
screen "EPROC-ALTAMS050" 1280x800, template "Plantilla-Alta-Sec"
   Button "Botón_3" at 467,294 size 40x38; TextOff 'Text'; PictureOff "x"
      on Click: function_efd93a16()
   Button "Botón_4" at 411,540 size 96x35; TextOff 'Hecho'; Authorization "Administración de usuarios"
      on Press: SetTag("Varios_UltimoMantMS050", "HorasSecAlta_HMMS050")
   TextField "Campo de texto_6" at 37,450 size 326x27; Text 'Tiempo de funcionamiento acumulado'
   TextField "Campo de texto_4" at 37,510 size 201x27; Text 'Próximo mantenimiento'
   IOField "Campo ES_7" at 25,475 size 173x35; Authorization "Administración de usuarios"; FormatPattern 999999999; Unit  hs
      ProcessValue <- "HorasSecAlta_HMMS050"
      Appearance <- "LimiteMantMS050"
   IOField "Campo ES_1" at 205,475 size 80x35; Authorization "Administración de usuarios"; FormatPattern 99; Unit  min
      ProcessValue <- "HorasSecAlta_MMMS050"
   IOField "Campo ES_2" at 25,535 size 173x35; FormatPattern 999999999; Unit  hs
      ProcessValue <- "ProxMantMS050"
      Appearance <- "LimiteMantMS050"
   GraphicIOField "Campo ES gráfico_3" at 21,434 size 511x6; PictureList "Indicador"
      ProcessValue <- "AnimaMS050"
   TextField "Campo de texto_3" at 46,356 size 89x39; Text 'ABC 1'
   SymbolicIOField "Campo ES simbólico_3" at 48,392 size 242x21; TextOff '0'; TextOn '1'; TextList "EstadoMotor"
      ProcessValue <- "AnimaMS050"
   Switch "Interruptor_8" at 205,359 size 29x29; TextOn '1'; TextOff '0'; CaptionText 'Switch'; PictureOff "A2"; Authorization "Operación"; PictureOn "A"
      ProcessValue <- "AutoMS050"
      Visibility <- "MantMS050"
   ScreenModuleView "Faceplate_2_4" at 274,346 size 244x69
      Guid_{11997190-23979} <- "HabilitaciónMS050"
      Guid_{11997190-37146} <- "Enc1MS050"
      Guid_{11997190-23983} <- "ParadaMS050"
      Guid_{11997190-23981} <- "MarchaMS050"
      Guid_{11997190-37150} <- "Enc2MS050"
      Guid_{11997190-23976} <- "DeshabilitaciónMS050"
      Guid_{11997190-23985} <- "AnimaMenuMS050"

screen "EPROC-ALTAMS051" 1280x800, template "Plantilla-Alta-Sec"
   Button "Botón_3" at 467,294 size 40x38; TextOff 'Text'; PictureOff "x"
      on Click: function_efd93a16()
   Button "Botón_4" at 411,540 size 96x35; TextOff 'Hecho'; Authorization "Administración de usuarios"
      on Press: SetTag("Varios_UltimoMantMS051", "HorasSecAlta_HMMS051")
   TextField "Campo de texto_6" at 37,450 size 326x27; Text 'Tiempo de funcionamiento acumulado'
   TextField "Campo de texto_4" at 37,510 size 201x27; Text 'Próximo mantenimiento'
   IOField "Campo ES_7" at 25,475 size 173x35; Authorization "Administración de usuarios"; FormatPattern 999999999; Unit  hs
      ProcessValue <- "HorasSecAlta_HMMS051"
      Appearance <- "LimiteMantMS051"
   IOField "Campo ES_1" at 205,475 size 80x35; Authorization "Administración de usuarios"; FormatPattern 99; Unit  min
      ProcessValue <- "HorasSecAlta_MMMS051"
   IOField "Campo ES_2" at 25,535 size 173x35; FormatPattern 999999999; Unit  hs
      ProcessValue <- "ProxMantMS051"
      Appearance <- "LimiteMantMS051"
   GraphicIOField "Campo ES gráfico_9" at 21,434 size 511x6; PictureList "Indicador"
      ProcessValue <- "AnimaMS051"
   TextField "Campo de texto_1" at 46,356 size 89x39; Text 'ABC 3'
   SymbolicIOField "Campo ES simbólico_9" at 48,392 size 242x21; TextOff '0'; TextOn '1'; TextList "EstadoMotor"
      ProcessValue <- "AnimaMS051"
   Switch "Interruptor_5" at 211,363 size 29x29; TextOn '1'; TextOff '0'; CaptionText 'Switch'; PictureOff "A2"; Authorization "Operación"; PictureOn "A"
      ProcessValue <- "AutoMS051"
      Visibility <- "MantMS051"
   ScreenModuleView "Faceplate_2_1" at 277,346 size 244x69
      Guid_{11997190-23979} <- "HabilitaciónMS051"
      Guid_{11997190-37146} <- "Enc1MS051"
      Guid_{11997190-23983} <- "ParadaMS051"
      Guid_{11997190-23981} <- "MarchaMS051"
      Guid_{11997190-37150} <- "Enc2MS051"
      Guid_{11997190-23976} <- "DeshabilitaciónMS051"
      Guid_{11997190-23985} <- "AnimaMenuMS051"

screen "EPROC-ALTAMS052" 1280x800, template "Plantilla-Alta-Sec"
   Button "Botón_3" at 467,294 size 40x38; TextOff 'Text'; PictureOff "x"
      on Click: function_efd93a16()
   Button "Botón_4" at 411,540 size 96x35; TextOff 'Hecho'; Authorization "Administración de usuarios"
      on Press: SetTag("Varios_UltimoMantMS052", "HorasSecAlta_HMMS052")
   TextField "Campo de texto_6" at 37,450 size 326x27; Text 'Tiempo de funcionamiento acumulado'
   TextField "Campo de texto_4" at 37,510 size 201x27; Text 'Próximo mantenimiento'
   IOField "Campo ES_7" at 25,475 size 173x35; Authorization "Administración de usuarios"; FormatPattern 999999999; Unit  hs
      ProcessValue <- "HorasSecAlta_HMMS052"
      Appearance <- "LimiteMantMS052"
   IOField "Campo ES_1" at 205,475 size 80x35; Authorization "Administración de usuarios"; FormatPattern 99; Unit  min
      ProcessValue <- "HorasSecAlta_MMMS052"
   IOField "Campo ES_2" at 25,535 size 173x35; FormatPattern 999999999; Unit  hs
      ProcessValue <- "ProxMantMS052"
      Appearance <- "LimiteMantMS052"
   GraphicIOField "Campo ES gráfico_1" at 21,434 size 511x6; PictureList "Indicador"
      ProcessValue <- "AnimaMS052"
   TextField "Campo de texto_1" at 46,356 size 89x39; Text 'ABC 2'
   SymbolicIOField "Campo ES simbólico_1" at 48,392 size 242x21; TextOff '0'; TextOn '1'; TextList "EstadoMotor"
      ProcessValue <- "AnimaMS052"
   Switch "Interruptor_6" at 227,365 size 29x29; TextOn '1'; TextOff '0'; CaptionText 'Switch'; PictureOff "A2"; Authorization "Operación"; PictureOn "A"
      ProcessValue <- "AutoMS052"
      Visibility <- "MantMS052"
   ScreenModuleView "Faceplate_2_2" at 277,346 size 244x69
      Guid_{11997190-23979} <- "HabilitaciónMS052"
      Guid_{11997190-37146} <- "Enc1MS052"
      Guid_{11997190-23983} <- "ParadaMS052"
      Guid_{11997190-23981} <- "MarchaMS052"
      Guid_{11997190-37150} <- "Enc2MS052"
      Guid_{11997190-23976} <- "DeshabilitaciónMS052"
      Guid_{11997190-23985} <- "AnimaMenuMS052"

screen "EPROC-ALTAMS053" 1280x800, template "Plantilla-Alta-Sec"
   Button "Botón_3" at 467,294 size 40x38; TextOff 'Text'; PictureOff "x"
      on Click: function_efd93a16()
   Button "Botón_4" at 411,540 size 96x35; TextOff 'Hecho'; Authorization "Administración de usuarios"
      on Press: SetTag("Varios_UltimoMantMS053", "HorasSecAlta_HMMS053")
   TextField "Campo de texto_6" at 37,450 size 326x27; Text 'Tiempo de funcionamiento acumulado'
   TextField "Campo de texto_4" at 37,510 size 201x27; Text 'Próximo mantenimiento'
   IOField "Campo ES_7" at 25,475 size 173x35; Authorization "Administración de usuarios"; FormatPattern 999999999; Unit  hs
      ProcessValue <- "HorasSecAlta_HMMS053"
      Appearance <- "LimiteMantMS053"
   IOField "Campo ES_1" at 205,475 size 80x35; Authorization "Administración de usuarios"; FormatPattern 99; Unit  min
      ProcessValue <- "HorasSecAlta_MMMS053"
   IOField "Campo ES_2" at 25,535 size 173x35; FormatPattern 999999999; Unit  hs
      ProcessValue <- "ProxMantMS053"
      Appearance <- "LimiteMantMS053"
   IOField "Campo ES_6" at 351,413 size 85x19; FormatPattern 999999999; Unit  hs
      ProcessValue <- "HorasSecAlta_HMMS053"
   GraphicIOField "Campo ES gráfico_2" at 21,434 size 511x6; PictureList "Indicador"
      ProcessValue <- "AnimaMS053"
   TextField "Campo de texto_2" at 46,351 size 101x39; Text 'Fargon'
   SymbolicIOField "Campo ES simbólico_2" at 48,387 size 242x21; TextOff '0'; TextOn '1'; TextList "EstadoMotor"
      ProcessValue <- "AnimaMS053"
   Switch "Interruptor_7" at 227,360 size 29x29; TextOn '1'; TextOff '0'; CaptionText 'Switch'; PictureOff "A2"; Authorization "Operación"; PictureOn "A"
      ProcessValue <- "AutoMS053"
      Visibility <- "MantMS053"
   ScreenModuleView "Faceplate_2_3" at 276,346 size 244x69
      Guid_{11997190-23979} <- "HabilitaciónMS053"
      Guid_{11997190-37146} <- "Enc1MS053"
      Guid_{11997190-23983} <- "ParadaMS053"
      Guid_{11997190-23981} <- "MarchaMS053"
      Guid_{11997190-37150} <- "Enc2MS053"
      Guid_{11997190-23976} <- "DeshabilitaciónMS053"
      Guid_{11997190-23985} <- "AnimaMenuMS053"

screen "EPROC-BAJAMC060" 1280x800, template "Plantilla-Baja-Cmp"
   Button "Botón_4" at 1135,405 size 96x35; TextOff 'Hecho'; Authorization "Administración de usuarios"
      on Press: SetTag("Varios_UltimoMantMC060_1", "HorasCmpBaja_HMMC060")
   TextField "Campo de texto_6" at 761,315 size 326x27; Text 'Tiempo de funcionamiento acumulado'
   TextField "Campo de texto_4" at 761,375 size 231x27; Text 'Próximo mantenimiento #1'
   Button "Botón_1" at 1135,470 size 96x35; TextOff 'Hecho'; Authorization "Administración de usuarios"
      on Press: SetTag("Varios_UltimoMantMC060_2", "HorasCmpBaja_HMMC060")
   TextField "Campo de texto_1" at 761,440 size 231x27; Text 'Próximo mantenimiento #2'
   Button "Botón_2" at 1135,535 size 96x35; TextOff 'Hecho'; Authorization "Administración de usuarios"
      on Press: SetTag("Varios_UltimoMantMC060_3", "HorasCmpBaja_HMMC060")
   TextField "Campo de texto_2" at 761,505 size 231x27; Text 'Próximo mantenimiento #3'
   Button "Botón_3" at 1135,600 size 96x35; TextOff 'Hecho'; Authorization "Administración de usuarios"
      on Press: SetTag("Varios_UltimoMantMC060_4", "HorasCmpBaja_HMMC060")
   TextField "Campo de texto_3" at 761,570 size 231x27; Text 'Próximo mantenimiento #4'
   Button "Botón_5" at 1135,665 size 96x35; TextOff 'Hecho'; Authorization "Administración de usuarios"
      on Press: SetTag("Varios_UltimoMantMC060_5", "HorasCmpBaja_HMMC060")
   TextField "Campo de texto_7" at 761,635 size 231x27; Text 'Próximo mantenimiento #5'
   Button "Botón_6" at 1199,168 size 40x38; TextOff 'Text'; PictureOff "x"
      on Click: function_efd93a16()
   GraphicIOField "Campo ES gráfico_4" at 746,294 size 511x6; PictureList "Indicador"
      ProcessValue <- "AnimaMC060"
   TextField "Campo de texto_5" at 771,224 size 116x39; Text 'Sullair 2'
   SymbolicIOField "Campo ES simbólico_9" at 773,260 size 242x21; TextOff '0'; TextOn '1'; TextList "EstadoMotor"
      ProcessValue <- "AnimaMC060"
   Switch "Interruptor_5" at 1108,242 size 91x31; TextOn 'Deshabilitado'; TextOff 'Habilitado'; CaptionText 'Switch'; Authorization "Administración de usuarios"
      Appearance <- "HabilitarMC060"
      ProcessValue <- "HabilitarMC060"
   IOField "Campo ES_7" at 749,340 size 173x35; Authorization "Administración de usuarios"; FormatPattern 999999999; Unit  hs
      ProcessValue <- "HorasCmpBaja_HMMC060"
      Appearance <- "EstadoMantMC060"
   IOField "Campo ES_1" at 929,340 size 80x35; Authorization "Administración de usuarios"; FormatPattern 99; Unit  min
      ProcessValue <- "HorasCmpBaja_MMMC060"
   IOField "Campo ES_2" at 749,400 size 173x35; FormatPattern 999999999; Unit  hs
      ProcessValue <- "ProxMantMC060_1"
      Appearance <- "LimiteMantMC060_1"
   IOField "Campo ES_3" at 749,465 size 173x35; FormatPattern 999999999; Unit  hs
      ProcessValue <- "ProxMantMC060_2"
      Appearance <- "LimiteMantMC060_2"
   IOField "Campo ES_4" at 749,530 size 173x35; FormatPattern 999999999; Unit  hs
      ProcessValue <- "ProxMantMC060_3"
      Appearance <- "LimiteMantMC060_3"
   IOField "Campo ES_5" at 749,595 size 173x35; FormatPattern 999999999; Unit  hs
      ProcessValue <- "ProxMantMC060_4"
      Appearance <- "LimiteMantMC060_4"
   IOField "Campo ES_6" at 749,660 size 173x35; FormatPattern 999999999; Unit  hs
      ProcessValue <- "ProxMantMC060_5"
      Appearance <- "LimiteMantMC060_5"

screen "EPROC-BAJAMC061" 1280x800, template "Plantilla-Baja-Cmp"
   Button "Botón_4" at 1135,405 size 96x35; TextOff 'Hecho'; Authorization "Administración de usuarios"
      on Press: SetTag("Varios_UltimoMantMC061_1", "HorasCmpBaja_HMMC061")
   TextField "Campo de texto_6" at 761,315 size 326x27; Text 'Tiempo de funcionamiento acumulado'
   TextField "Campo de texto_4" at 761,375 size 231x27; Text 'Próximo mantenimiento #1'
   Button "Botón_1" at 1135,470 size 96x35; TextOff 'Hecho'; Authorization "Administración de usuarios"
      on Press: SetTag("Varios_UltimoMantMC061_2", "HorasCmpBaja_HMMC061")
   TextField "Campo de texto_1" at 761,440 size 231x27; Text 'Próximo mantenimiento #2'
   Button "Botón_2" at 1135,535 size 96x35; TextOff 'Hecho'; Authorization "Administración de usuarios"
      on Press: SetTag("Varios_UltimoMantMC061_3", "HorasCmpBaja_HMMC061")
   TextField "Campo de texto_2" at 761,505 size 231x27; Text 'Próximo mantenimiento #3'
   Button "Botón_3" at 1135,600 size 96x35; TextOff 'Hecho'; Authorization "Administración de usuarios"
      on Press: SetTag("Varios_UltimoMantMC061_4", "HorasCmpBaja_HMMC061")
   TextField "Campo de texto_3" at 761,570 size 231x27; Text 'Próximo mantenimiento #4'
   Button "Botón_5" at 1135,665 size 96x35; TextOff 'Hecho'; Authorization "Administración de usuarios"
      on Press: SetTag("Varios_UltimoMantMC061_5", "HorasCmpBaja_HMMC061")
   TextField "Campo de texto_7" at 761,635 size 231x27; Text 'Próximo mantenimiento #5'
   Button "Botón_6" at 1199,168 size 40x38; TextOff 'Text'; PictureOff "x"
      on Click: function_efd93a16()
   IOField "Campo ES_7" at 749,340 size 173x35; Authorization "Administración de usuarios"; FormatPattern 999999999; Unit  hs
      ProcessValue <- "HorasCmpBaja_HMMC061"
      Appearance <- "EstadoMantMC061"
   IOField "Campo ES_1" at 929,340 size 80x35; Authorization "Administración de usuarios"; FormatPattern 99; Unit  min
      ProcessValue <- "HorasCmpBaja_MMMC061"
   IOField "Campo ES_2" at 749,400 size 173x35; FormatPattern 999999999; Unit  hs
      Appearance <- "LimiteMantMS051"
      ProcessValue <- "ProxMantMC061_1"
   IOField "Campo ES_3" at 749,465 size 173x35; FormatPattern 999999999; Unit  hs
      Appearance <- "LimiteMantMS051"
      ProcessValue <- "ProxMantMC061_2"
   IOField "Campo ES_4" at 749,530 size 173x35; FormatPattern 999999999; Unit  hs
      Appearance <- "LimiteMantMS051"
      ProcessValue <- "ProxMantMC061_3"
   IOField "Campo ES_5" at 749,595 size 173x35; FormatPattern 999999999; Unit  hs
      Appearance <- "LimiteMantMS051"
      ProcessValue <- "ProxMantMC061_4"
   IOField "Campo ES_6" at 749,660 size 173x35; FormatPattern 999999999; Unit  hs
      Appearance <- "LimiteMantMS051"
      ProcessValue <- "ProxMantMC061_5"
   GraphicIOField "Campo ES gráfico_3" at 746,293 size 510x6; PictureList "Indicador"
      ProcessValue <- "AnimaMC061"
   TextField "Campo de texto_5" at 771,224 size 116x39; Text 'Sullair 1'
   SymbolicIOField "Campo ES simbólico_8" at 773,260 size 242x21; TextOff '0'; TextOn '1'; TextList "EstadoMotor"
      ProcessValue <- "AnimaMC061"
   Switch "Interruptor_4" at 974,228 size 29x29; TextOn '1'; TextOff '0'; CaptionText 'Switch'; PictureOff "A2"; Authorization "Operación"; PictureOn "A"
      ProcessValue <- "AutoMC061"
      Visibility <- "MantM061"
   ScreenModuleView "Faceplate_1_1" at 1018,228 size 236x58
      Guid_{11997190-23979} <- "HabilitaciónMC061"
      Guid_{11997190-23983} <- "ParadaMC061"
      Guid_{11997190-23981} <- "MarchaMC061"
      Guid_{11997190-23989} <- "SpoffMC061"
      Guid_{11997190-23976} <- "DeshabilitaciónMC061"
      Guid_{11997190-23987} <- "SponMC061"
      Guid_{11997190-23985} <- "AnimMenuMC061"

screen "EPROC-BAJAMC062" 1280x800, template "Plantilla-Baja-Cmp"
   Button "Botón_4" at 1135,405 size 96x35; TextOff 'Hecho'; Authorization "Administración de usuarios"
      on Press: SetTag("Varios_UltimoMantMC062_1", "HorasCmpBaja_HMMC062")
   TextField "Campo de texto_6" at 761,315 size 326x27; Text 'Tiempo de funcionamiento acumulado'
   TextField "Campo de texto_4" at 761,375 size 231x27; Text 'Próximo mantenimiento #1'
   Button "Botón_1" at 1135,470 size 96x35; TextOff 'Hecho'; Authorization "Administración de usuarios"
      on Press: SetTag("Varios_UltimoMantMC062_2", "HorasCmpBaja_HMMC062")
   TextField "Campo de texto_1" at 761,440 size 231x27; Text 'Próximo mantenimiento #2'
   Button "Botón_2" at 1135,535 size 96x35; TextOff 'Hecho'; Authorization "Administración de usuarios"
      on Press: SetTag("Varios_UltimoMantMC062_3", "HorasCmpBaja_HMMC062")
   TextField "Campo de texto_2" at 761,505 size 231x27; Text 'Próximo mantenimiento #3'
   Button "Botón_3" at 1135,600 size 96x35; TextOff 'Hecho'; Authorization "Administración de usuarios"
      on Press: SetTag("Varios_HorasMantMC062_4", "HorasCmpBaja_HMMC062")
   TextField "Campo de texto_3" at 761,570 size 231x27; Text 'Próximo mantenimiento #4'
   Button "Botón_5" at 1135,665 size 96x35; TextOff 'Hecho'; Authorization "Administración de usuarios"
      on Press: SetTag("Varios_UltimoMantMC062_5", "HorasCmpBaja_HMMC062")
   TextField "Campo de texto_7" at 761,635 size 231x27; Text 'Próximo mantenimiento #5'
   Button "Botón_6" at 1199,168 size 40x38; TextOff 'Text'; PictureOff "x"
      on Click: function_efd93a16()
   IOField "Campo ES_7" at 749,340 size 173x35; Authorization "Administración de usuarios"; FormatPattern 999999999; Unit  hs
      ProcessValue <- "HorasCmpBaja_HMMC062"
      Appearance <- "EstadoMantMC062"
   IOField "Campo ES_1" at 929,340 size 80x35; Authorization "Administración de usuarios"; FormatPattern 99; Unit  min
      ProcessValue <- "HorasCmpBaja_MMMC062"
   IOField "Campo ES_2" at 749,400 size 173x35; FormatPattern 999999999; Unit  hs
      Appearance <- "LimiteMantMS051"
      ProcessValue <- "ProxMantMC062_1"
   IOField "Campo ES_3" at 749,465 size 173x35; FormatPattern 999999999; Unit  hs
      Appearance <- "LimiteMantMS051"
      ProcessValue <- "ProxMantMC062_2"
   IOField "Campo ES_4" at 749,530 size 173x35; FormatPattern 999999999; Unit  hs
      Appearance <- "LimiteMantMS051"
      ProcessValue <- "ProxMantMC062_3"
   IOField "Campo ES_5" at 749,595 size 173x35; FormatPattern 999999999; Unit  hs
      Appearance <- "LimiteMantMS051"
      ProcessValue <- "ProxMantMC062_4"
   IOField "Campo ES_6" at 749,660 size 173x35; FormatPattern 999999999; Unit  hs
      Appearance <- "LimiteMantMS051"
      ProcessValue <- "ProxMantMC062_5"
   GraphicIOField "Campo ES gráfico_2" at 747,293 size 507x6; PictureList "Indicador"
      ProcessValue <- "AnimaMC062"
   TextField "Campo de texto_5" at 771,224 size 116x39; Text 'Sullair 0'
   SymbolicIOField "Campo ES simbólico_7" at 773,260 size 242x21; TextOff '0'; TextOn '1'; TextList "EstadoMotor"
      ProcessValue <- "AnimaMC062"
   Switch "Interruptor_3" at 970,227 size 29x29; TextOn '1'; TextOff '0'; CaptionText 'Switch'; PictureOff "A2"; Authorization "Operación"; PictureOn "A"
      ProcessValue <- "AutoMC062"
      Visibility <- "MantM062"
   ScreenModuleView "Faceplate_1_3" at 1013,227 size 236x58
      Guid_{11997190-23979} <- "HabilitaciónMC062"
      Guid_{11997190-23983} <- "ParadaMC062"
      Guid_{11997190-23981} <- "MarchaMC062"
      Guid_{11997190-23989} <- "SpoffMC062"
      Guid_{11997190-23976} <- "DeshabilitaciónMC062"
      Guid_{11997190-23987} <- "SponMC062"
      Guid_{11997190-23985} <- "AnimMenuMC062"

screen "EPROC-BAJAMC063" 1280x800, template "Plantilla-Baja-Cmp"
   Button "Botón_4" at 1135,405 size 96x35; TextOff 'Hecho'; Authorization "Administración de usuarios"
      on Press: SetTag("Varios_UltimoMantMC063_1", "HorasCmpBaja_HMMC063")
   TextField "Campo de texto_6" at 761,315 size 326x27; Text 'Tiempo de funcionamiento acumulado'
   TextField "Campo de texto_4" at 761,375 size 231x27; Text 'Próximo mantenimiento #1'
   Button "Botón_1" at 1135,470 size 96x35; TextOff 'Hecho'; Authorization "Administración de usuarios"
      on Press: SetTag("Varios_UltimoMantMC063_2", "HorasCmpBaja_HMMC063")
   TextField "Campo de texto_1" at 761,440 size 231x27; Text 'Próximo mantenimiento #2'
   Button "Botón_2" at 1135,535 size 96x35; TextOff 'Hecho'; Authorization "Administración de usuarios"
      on Press: SetTag("Varios_UltimoMantMC063_3", "HorasCmpBaja_HMMC063")
   TextField "Campo de texto_2" at 761,505 size 231x27; Text 'Próximo mantenimiento #3'
   Button "Botón_3" at 1135,600 size 96x35; TextOff 'Hecho'; Authorization "Administración de usuarios"
      on Press: SetTag("Varios_UltimoMantMC063_4", "HorasCmpBaja_HMMC063")
   TextField "Campo de texto_3" at 761,570 size 231x27; Text 'Próximo mantenimiento #4'
   Button "Botón_5" at 1135,665 size 96x35; TextOff 'Hecho'; Authorization "Administración de usuarios"
      on Press: SetTag("Varios_UltimoMantMC063_5", "HorasCmpBaja_HMMC063")
   TextField "Campo de texto_7" at 761,635 size 231x27; Text 'Próximo mantenimiento #5'
   Button "Botón_6" at 1199,168 size 40x38; TextOff 'Text'; PictureOff "x"
      on Click: function_efd93a16()
   IOField "Campo ES_7" at 749,340 size 173x35; Authorization "Administración de usuarios"; FormatPattern 999999999; Unit  hs
      ProcessValue <- "HorasCmpBaja_HMMC063"
      Appearance <- "EstadoMantMC063"
   IOField "Campo ES_1" at 929,340 size 80x35; Authorization "Administración de usuarios"; FormatPattern 99; Unit  min
      ProcessValue <- "HorasCmpBaja_MMMC063"
   IOField "Campo ES_2" at 749,400 size 173x35; FormatPattern 999999999; Unit  hs
      Appearance <- "LimiteMantMS051"
      ProcessValue <- "ProxMantMC063_1"
   IOField "Campo ES_3" at 749,465 size 173x35; FormatPattern 999999999; Unit  hs
      Appearance <- "LimiteMantMS051"
      ProcessValue <- "ProxMantMC063_2"
   IOField "Campo ES_4" at 749,530 size 173x35; FormatPattern 999999999; Unit  hs
      Appearance <- "LimiteMantMS051"
      ProcessValue <- "ProxMantMC063_3"
   IOField "Campo ES_5" at 749,595 size 173x35; FormatPattern 999999999; Unit  hs
      Appearance <- "LimiteMantMS051"
      ProcessValue <- "ProxMantMC063_4"
   IOField "Campo ES_6" at 749,660 size 173x35; FormatPattern 999999999; Unit  hs
      Appearance <- "LimiteMantMS051"
      ProcessValue <- "ProxMantMC063_5"
   GraphicIOField "Campo ES gráfico_1" at 746,293 size 507x6; PictureList "Indicador"
      ProcessValue <- "AnimaMC063"
   TextField "Campo de texto_8" at 763,224 size 91x39; Text 'Atlas 3'
   SymbolicIOField "Campo ES simbólico_6" at 765,260 size 242x21; TextOff '0'; TextOn '1'; TextList "EstadoMotor"
      ProcessValue <- "AnimaMC063"
   Switch "Interruptor_2" at 967,227 size 29x29; TextOn '1'; TextOff '0'; CaptionText 'Switch'; PictureOff "A2"; Authorization "Operación"; PictureOn "A"
      ProcessValue <- "AutoMC063"
      Visibility <- "MantM063"
   ScreenModuleView "Faceplate_1_4" at 1014,226 size 236x58
      Guid_{11997190-23979} <- "HabilitaciónMC063"
      Guid_{11997190-23983} <- "ParadaMC063"
      Guid_{11997190-23981} <- "MarchaMC063"
      Guid_{11997190-23989} <- "SpoffMC063"
      Guid_{11997190-23976} <- "DeshabilitaciónMC063"
      Guid_{11997190-23987} <- "SponMC063"
      Guid_{11997190-23985} <- "AnimMenuMC063"

screen "EPROC-BAJAMC064" 1280x800, template "Plantilla-Baja-Cmp"
   Button "Botón_4" at 1135,405 size 96x35; TextOff 'Hecho'; Authorization "Administración de usuarios"
      on Press: SetTag("Varios_UltimoMantMC064_1", "HorasCmpBaja_HMMC064")
   TextField "Campo de texto_6" at 761,315 size 326x27; Text 'Tiempo de funcionamiento acumulado'
   TextField "Campo de texto_4" at 761,375 size 231x27; Text 'Próximo mantenimiento #1'
   Button "Botón_1" at 1135,470 size 96x35; TextOff 'Hecho'; Authorization "Administración de usuarios"
      on Press: SetTag("Varios_UltimoMantMC064_2", "HorasCmpBaja_HMMC064")
   TextField "Campo de texto_1" at 761,440 size 231x27; Text 'Próximo mantenimiento #2'
   Button "Botón_2" at 1135,535 size 96x35; TextOff 'Hecho'; Authorization "Administración de usuarios"
      on Press: SetTag("Varios_UltimoMantMC064_3", "HorasCmpBaja_HMMC064")
   TextField "Campo de texto_2" at 761,505 size 231x27; Text 'Próximo mantenimiento #3'
   Button "Botón_3" at 1135,600 size 96x35; TextOff 'Hecho'; Authorization "Administración de usuarios"
      on Press: SetTag("Varios_UltimoMantMC064_4", "HorasCmpBaja_HMMC064")
   TextField "Campo de texto_3" at 761,570 size 231x27; Text 'Próximo mantenimiento #4'
   Button "Botón_5" at 1135,665 size 96x35; TextOff 'Hecho'; Authorization "Administración de usuarios"
      on Press: SetTag("Varios_UltimoMantMC064_5", "HorasCmpBaja_HMMC064")
   TextField "Campo de texto_7" at 761,635 size 231x27; Text 'Próximo mantenimiento #5'
   Button "Botón_6" at 1199,168 size 40x38; TextOff 'Text'; PictureOff "x"
      on Click: function_efd93a16()
   IOField "Campo ES_7" at 749,340 size 173x35; Authorization "Administración de usuarios"; FormatPattern 999999999; Unit  hs
      ProcessValue <- "HorasCmpBaja_HMMC064"
      Appearance <- "EstadoMantMC064"
   IOField "Campo ES_1" at 929,340 size 80x35; Authorization "Administración de usuarios"; FormatPattern 99; Unit  min
      ProcessValue <- "HorasCmpBaja_MMMC064"
   IOField "Campo ES_2" at 749,400 size 173x35; FormatPattern 999999999; Unit  hs
      Appearance <- "LimiteMantMS051"
      ProcessValue <- "ProxMantMC064_1"
   IOField "Campo ES_3" at 749,465 size 173x35; FormatPattern 999999999; Unit  hs
      Appearance <- "LimiteMantMS051"
      ProcessValue <- "ProxMantMC064_2"
   IOField "Campo ES_4" at 749,530 size 173x35; FormatPattern 999999999; Unit  hs
      Appearance <- "LimiteMantMS051"
      ProcessValue <- "ProxMantMC064_3"
   IOField "Campo ES_5" at 749,595 size 173x35; FormatPattern 999999999; Unit  hs
      Appearance <- "LimiteMantMS051"
      ProcessValue <- "ProxMantMC064_4"
   IOField "Campo ES_6" at 749,660 size 173x35; FormatPattern 999999999; Unit  hs
      Appearance <- "LimiteMantMS051"
      ProcessValue <- "ProxMantMC064_5"
   GraphicIOField "Campo ES gráfico_5" at 747,294 size 507x6; PictureList "Indicador"
      ProcessValue <- "AnimaMC064"
   TextField "Campo de texto_9" at 771,224 size 100x39; Text 'Atlas 2'
   SymbolicIOField "Campo ES simbólico_5" at 773,260 size 242x21; TextOff '0'; TextOn '1'; TextList "EstadoMotor"
      ProcessValue <- "AnimaMC064"
   Switch "Interruptor_1" at 969,227 size 29x29; TextOn '1'; TextOff '0'; CaptionText 'Switch'; PictureOff "A2"; Authorization "Operación"; PictureOn "A"
      ProcessValue <- "AutoMC064"
      Visibility <- "MantM064"
   ScreenModuleView "Faceplate_1_5" at 1016,227 size 236x58
      Guid_{11997190-23979} <- "HabilitaciónMC064"
      Guid_{11997190-23983} <- "ParadaMC064"
      Guid_{11997190-23981} <- "MarchaMC064"
      Guid_{11997190-23989} <- "SpoffMC064"
      Guid_{11997190-23976} <- "DeshabilitaciónMC064"
      Guid_{11997190-23987} <- "SponMC064"
      Guid_{11997190-23985} <- "AnimMenuMC064"

screen "EPROC-BAJAMS054" 1280x800, template "Plantilla-Baja-Sec"
   TextField "Campo de texto_1" at 758,509 size 326x27; Text 'Tiempo de funcionamiento acumulado'
   Button "Botón_4" at 1032,599 size 96x35; TextOff 'Hecho'; Authorization "Administración de usuarios"
      on Press: SetTag("Varios_UltimoMantMS054_1", "HorasSecBaja_HMMS054")
   TextField "Campo de texto_4" at 758,569 size 231x27; Text 'Próximo mantenimiento #1'
   TextField "Campo de texto_5" at 758,634 size 231x27; Text 'Próximo mantenimiento #2'
   Button "Botón_5" at 1032,664 size 96x35; TextOff 'Hecho'; Authorization "Administración de usuarios"
      on Press: SetTag("Varios_UltimoMantMS054_2", "HorasSecBaja_HMMS054")
   Button "Botón_6" at 1188,358 size 40x38; TextOff 'Text'; PictureOff "x"
      on Click: function_efd93a16()
   IOField "Campo ES_7" at 746,534 size 173x35; Authorization "Administración de usuarios"; FormatPattern 999999999; Unit  hs
      ProcessValue <- "HorasSecBaja_HMMS054"
      Appearance <- "EstadoMantSecBaja"
   IOField "Campo ES_1" at 926,534 size 80x35; Authorization "Administración de usuarios"; FormatPattern 99; Unit  min
      ProcessValue <- "HorasSecBaja_MMMS054"
   IOField "Campo ES_2" at 746,594 size 173x35; FormatPattern 999999999; Unit  hs
      ProcessValue <- "ProxMantMS054_1"
      Appearance <- "LimiteMantMS054_1"
   IOField "Campo ES_3" at 746,659 size 173x35; FormatPattern 999999999; Unit  hs
      ProcessValue <- "ProxMantMS054_2"
      Appearance <- "LimiteMantMS054_2"
   GraphicIOField "Campo ES gráfico_3" at 736,489 size 510x6; PictureList "Indicador"
      ProcessValue <- "AnimaMS054"
   TextField "Campo de texto_6" at 761,411 size 116x39; Text 'Sullair 1'
   SymbolicIOField "Campo ES simbólico_8" at 763,447 size 242x21; TextOff '0'; TextOn '1'; TextList "EstadoMotor"
      ProcessValue <- "AnimaMS054"
   ScreenModuleView "Faceplate_3_1" at 1015,411 size 213x73; ScreenModuleType ""
      Guid_{11997190-23981} <- "MarchaMS054"
      Guid_{11997190-23979} <- "HabilitaciónMS054"
      Guid_{11997190-23976} <- "DeshabilitaciónMS054"
      Guid_{11997190-23983} <- "ParadaMS054"

screen "EPROC-BAJAMS055" 1280x800, template "Plantilla-Baja-Sec"
   TextField "Campo de texto_1" at 758,509 size 326x27; Text 'Tiempo de funcionamiento acumulado'
   Button "Botón_4" at 1032,599 size 96x35; TextOff 'Hecho'; Authorization "Administración de usuarios"
      on Press: SetTag("Varios_UltimoMantMS055_1", "HorasSecBaja_HMMS055")
   TextField "Campo de texto_4" at 758,569 size 231x27; Text 'Próximo mantenimiento #1'
   TextField "Campo de texto_5" at 758,634 size 231x27; Text 'Próximo mantenimiento #2'
   Button "Botón_5" at 1032,664 size 96x35; TextOff 'Hecho'; Authorization "Administración de usuarios"
      on Press: SetTag("Varios_UltimoMantMS055_2", "HorasSecBaja_HMMS055")
   Button "Botón_6" at 1188,358 size 40x38; TextOff 'Text'; PictureOff "x"
      on Click: function_efd93a16()
   IOField "Campo ES_7" at 746,534 size 173x35; Authorization "Administración de usuarios"; FormatPattern 999999999; Unit  hs
      Appearance <- "EstadoMantSecBaja"
      ProcessValue <- "HorasSecBaja_HMMS055"
   IOField "Campo ES_1" at 926,534 size 80x35; Authorization "Administración de usuarios"; FormatPattern 99; Unit  min
      ProcessValue <- "HorasSecBaja_MMMS055"
   IOField "Campo ES_2" at 746,594 size 173x35; FormatPattern 999999999; Unit  hs
      Appearance <- "LimiteMantMS055_1"
      ProcessValue <- "ProxMantMS055_1"
   IOField "Campo ES_3" at 746,659 size 173x35; FormatPattern 999999999; Unit  hs
      Appearance <- "LimiteMantMS055_2"
      ProcessValue <- "ProxMantMS055_2"
   GraphicIOField "Campo ES gráfico_4" at 736,489 size 511x6; PictureList "Indicador"
      ProcessValue <- "AnimaMS055"
   TextField "Campo de texto_2" at 761,411 size 116x39; Text 'Sullair 2'
   SymbolicIOField "Campo ES simbólico_9" at 763,447 size 242x21; TextOff '0'; TextOn '1'; TextList "EstadoMotor"
      ProcessValue <- "AnimaMS055"
   ScreenModuleView "Faceplate_3_2" at 1020,411 size 213x73; ScreenModuleType ""
      Guid_{11997190-23981} <- "MarchaMS055"
      Guid_{11997190-23979} <- "HabilitaciónMS055"
      Guid_{11997190-23976} <- "DeshabilitaciónMS055"
      Guid_{11997190-23983} <- "ParadaMS055"

screen "Imagen_1" 1280x800
   GraphicIOField "Campo ES gráfico_3" at 736,489 size 510x6; PictureList "Indicador"
      ProcessValue <- "AnimaMS054"
   TextField "Campo de texto_6" at 761,411 size 116x39; Text 'Sullair 1'
   SymbolicIOField "Campo ES simbólico_8" at 763,447 size 242x21; TextOff '0'; TextOn '1'; TextList "EstadoMotor"
      ProcessValue <- "AnimaMS054"
   ScreenModuleView "Faceplate_3_1" at 1015,411 size 213x73; ScreenModuleType ""
      Guid_{11997190-23981} <- "MarchaMS054"
      Guid_{11997190-23979} <- "HabilitaciónMS054"
      Guid_{11997190-23976} <- "DeshabilitaciónMS054"
      Guid_{11997190-23983} <- "ParadaMS054"

Template "Plantilla" 1280x800
   Button "Plantilla_6" at 1196,741 size 81x58; TextOff 'Reconocer'; PictureOff "Asleep Check Mark Icon - Sleep Aid Records_2"
      on Press: SetBit("ReconocerTODAS")
      on Release: ResetBit("ReconocerTODAS")
      Appearance <- "AlarmaNueva"
   Button "Plantilla_1" at 1037,749 size 78x50; TextOff 'Anular Sirena'
      on Click: SetBit("AnularSirena?")
   Button "Plantilla_3" at 717,748 size 78x50; TextOff 'Text'; PictureOff "Rayo"
      on Click: ActivateScreen("SentronPAC-MTA", 0)
   Button "Plantilla_4" at 877,748 size 78x50; TextOff 'Text'
   Button "Plantilla_5" at 957,748 size 78x50; TextOff 'Parar Runtime'
      on Click: StopRuntime(0)
   Button "Plantilla_7" at 479,748 size 78x50; TextOff 'Compres.'
      on Click: ActivateScreen("MTA-CompBAJA", 0)
   Button "Plantilla_8" at 161,748 size 78x50; TextOff 'Torres'
      on Release: ActivateScreen("MTA-TorresCH", 0)
   Button "Plantilla_9" at 81,748 size 78x50; TextOff 'General'; TextOn 'NavigateHome'; PictureOff "NavigateHome_HMI_1"; PictureOn "NavigateHome_HMI_1"
      on Press: ResetBit("VerCh1MTA"); ResetBit("VerCh2MTA"); ResetBit("VerCh3MTA"); ResetBit("VerCh4MTA")
      on Release: ActivateScreen("MTA-Chillers-General", 0)
   Button "Plantilla_10" at 1117,741 size 78x58; TextOff 'Avisos'
      on Click: ActivateScreen("MTA-Avisos", 0)
      Appearance <- "AlarmaNueva"
   Button "Plantilla_12" at 638,748 size 78x50; TextOff 'Luz'; PictureOff "Lamp2_1"
      on Click: ActivateScreen("IluminaciónMTA", 0)
      Appearance <- "MantenerON"
   Button "Plantilla_13" at 400,748 size 78x50; TextOff 'Torres'
      on Click: ActivateScreen("MTA-TorresCAV", 0)
   Button "Plantilla_14" at 321,748 size 78x50; TextOff 'Secadores'
      on Click: ActivateScreen("MTA-SecALTA", 0)
   Button "Plantilla_15" at 558,748 size 78x50; TextOff 'Secadores'
      on Click: ActivateScreen("MTA-SecBaja", 0)
   Button "Plantilla_16" at 241,748 size 78x50; TextOff 'Compres.'
      on Click: ActivateScreen("MTA-CompALTA", 0)
   Button "Plantilla_17" at 1,740 size 78x58; TextOff 'NavigateHome'; PictureOff "NavigateHome_HMI_1"; PictureOn "NavigateHome_HMI_1"
      on Release: ActivateScreen("INICIO", 0)
   GraphicView "Plantilla_Visor de gráficos_1" at 80,740 size 78x6; Picture "indGris"
   GraphicView "Plantilla_Visor de gráficos_2" at 160,740 size 78x6; Picture "indGris"
   GraphicView "Plantilla_Visor de gráficos_3" at 478,740 size 78x6; Picture "indGris"
   GraphicView "Plantilla_Visor de gráficos_4" at 240,740 size 78x6; Picture "indGris"
   GraphicView "Plantilla_Visor de gráficos_5" at 557,740 size 78x6; Picture "indGris"
   GraphicView "Plantilla_Visor de gráficos_6" at 320,740 size 78x6; Picture "indGris"
   GraphicView "Plantilla_Visor de gráficos_7" at 399,740 size 78x6; Picture "indGris"
   GraphicView "Plantilla_Visor de gráficos_11" at 637,740 size 78x6; Picture "indGris"
   GraphicView "Plantilla_Visor de gráficos_8" at 80,740 size 78x6; Picture "indAmarillo"
      Visibility <- "IndCh"
   GraphicView "Plantilla_Visor de gráficos_9" at 160,740 size 78x6; Picture "indAmarillo"
      Visibility <- "IndTrCh"
   GraphicView "Plantilla_Visor de gráficos_10" at 478,740 size 78x6; Picture "indAmarillo"
      Visibility <- "IndCmpBaja"
   GraphicView "Plantilla_Visor de gráficos_12" at 240,740 size 78x6; Picture "indAmarillo"
      Visibility <- "IndCmpAlta"
   GraphicView "Plantilla_Visor de gráficos_13" at 557,740 size 78x6; Picture "indAmarillo"
      Visibility <- "IndSecBaja"
   GraphicView "Plantilla_Visor de gráficos_14" at 320,740 size 78x6; Picture "indAmarillo"
      Visibility <- "IndSecAlta"
   GraphicView "Plantilla_Visor de gráficos_15" at 399,740 size 78x6; Picture "indAmarillo"
      Visibility <- "IndTrCav"
   GraphicView "Plantilla_Visor de gráficos_16" at 637,740 size 78x6; Picture "indAmarillo"
      Visibility <- "MantenerON"
   TextField "Plantilla_Campo de texto_2" at 521,711 size 69x18; Text 'Baja Presión'
   TextField "Plantilla_Campo de texto_4" at 323,711 size 68x18; Text 'Alta Presión'
   TextField "Plantilla_Campo de texto_1" at 139,711 size 40x18; Text 'Chillers'
   Button "Plantilla_11" at 797,748 size 78x50; TextOff 'Variables Analóg.'
      on Click: ActivateScreen("Grafica", 0)
   GraphicView "Plantilla_Visor de gráficos_18" at 717,740 size 78x6; Picture "indGris"
   GraphicView "Plantilla_Visor de gráficos_19" at 797,740 size 78x6; Picture "indGris"
   GraphicView "Plantilla_Visor de gráficos_20" at 877,740 size 78x6; Picture "indGris"
   GraphicView "Plantilla_Visor de gráficos_21" at 957,740 size 78x6; Picture "indGris"
   GraphicView "Plantilla_Visor de gráficos_22" at 1037,741 size 78x6; Picture "indGris"
   GraphicView "Plantilla_Visor de gráficos_23" at 1037,741 size 78x6; Picture "indAmarillo"
      Visibility <- "AnularSirenaCav"
   GraphicView "Plantilla_Visor de gráficos_24" at 877,740 size 78x6; Picture "indAmarillo"
      Visibility <- "AlarmaBoosters"
   Group "Group" at 3,716 size 1276x83
   GraphicView "Plantilla_Visor de gráficos_26" at 68,9 size 91x26; Picture "eProC logo 4 b"
   GraphicView "Plantilla_Visor de gráficos_27" at 9,8 size 49x29; Picture "eProC logo 4 a"
   Rectangle "Plantilla_Rectángulo_1" at 3,716 size 1276x83
      Visibility <- "AnularSirena?"
   TextField "Plantilla_Campo de texto_3" at 34,732 size 696x50; Text '¿Está seguro de ANULAR la sirena? Si decide anular el sistema dejará de emitir avisos sonoros de manera permanente'
      Visibility <- "AnularSirena?"
   Button "Plantilla_Botón_1" at 1234,724 size 37x34; TextOff 'x'
      on Click: ResetBit("AnularSirena?")
      Visibility <- "AnularSirena?"
   Button "Plantilla_Botón_2" at 947,735 size 112x46; TextOff 'Activar'
      on Click: ResetBit("AnularSirenaCav")
      Visibility <- "AnularSirena?"
      Appearance <- "AnularSirenaCav"
   Button "Plantilla_Botón_3" at 1067,735 size 112x46; TextOff 'Desactivar'
      on Click: SetBit("AnularSirenaCav")
      Visibility <- "AnularSirena?"
      Appearance <- "AnularSirenaCav"

Template "Plantilla-Alta-Cmp" 1280x800
   Rectangle "Plantilla_Rectángulo_1" at 1,716 size 1276x84
      Visibility <- "AnularSirena?"
   TextField "Plantilla_Campo de texto_5" at 32,732 size 696x50; Text '¿Está seguro de ANULAR la sirena? Si decide anular el sistema dejará de emitir avisos sonoros de manera permanente'
      Visibility <- "AnularSirena?"
   Button "Plantilla_Botón_1" at 1232,724 size 37x34; TextOff 'x'
      on Click: ResetBit("AnularSirena?")
      Visibility <- "AnularSirena?"
   Button "Plantilla_Botón_2" at 945,735 size 112x46; TextOff 'Activar'
      on Click: ResetBit("AnularSirenaCav")
      Visibility <- "AnularSirena?"
      Appearance <- "AnularSirenaCav"
   Button "Plantilla_Botón_3" at 1065,735 size 112x46; TextOff 'Desactivar'
      on Click: SetBit("AnularSirenaCav")
      Visibility <- "AnularSirena?"
      Appearance <- "AnularSirenaCav"
   GraphicView "Visor de gráficos_8" at 1175,577 size 29x50; Picture "Gráfico_2"
   GraphicView "Visor de gráficos_7" at 885,605 size 391x113; Picture "tanque1X2"
   Button "Plantilla_6" at 1196,741 size 81x58; TextOff 'Reconocer'; PictureOff "Asleep Check Mark Icon - Sleep Aid Records_2"
      on Press: SetBit("ReconocerTODAS")
      on Release: ResetBit("ReconocerTODAS")
      Appearance <- "AlarmaNueva"
   GraphicView "Plantilla_Visor de gráficos_17" at 4,4 size 87x38; Picture "logo4"
   Button "Plantilla_7" at 479,748 size 78x50; TextOff 'Compres.'
      on Click: ActivateScreen("MTA-CompBAJA", 0)
   Button "Plantilla_8" at 161,748 size 78x50; TextOff 'Torres'
      on Release: ActivateScreen("MTA-TorresCH", 0)
   Button "Plantilla_9" at 81,748 size 78x50; TextOff 'General'; TextOn 'NavigateHome'; PictureOff "NavigateHome_HMI_1"; PictureOn "NavigateHome_HMI_1"
      on Press: ResetBit("VerCh1MTA"); ResetBit("VerCh2MTA"); ResetBit("VerCh3MTA"); ResetBit("VerCh4MTA")
      on Release: ActivateScreen("MTA-Chillers-General", 0)
   Button "Plantilla_12" at 638,748 size 78x50; TextOff 'Luz'; PictureOff "Lamp2_1"
      on Click: ActivateScreen("IluminaciónMTA", 0)
      Appearance <- "MantenerON"
   Button "Plantilla_13" at 400,748 size 78x50; TextOff 'Torres'
      on Click: ActivateScreen("MTA-TorresCAV", 0)
   Button "Plantilla_14" at 321,748 size 78x50; TextOff 'Secadores'
      on Click: ActivateScreen("MTA-SecALTA", 0)
   Button "Plantilla_15" at 558,748 size 78x50; TextOff 'Secadores'
      on Click: ActivateScreen("MTA-SecBaja", 0)
   Button "Plantilla_16" at 241,748 size 78x50; TextOff 'Compres.'
      on Click: ActivateScreen("MTA-CompALTA", 0)
   Button "Plantilla_17" at 1,740 size 78x58; TextOff 'NavigateHome'; PictureOff "NavigateHome_HMI_1"; PictureOn "NavigateHome_HMI_1"
      on Release: ActivateScreen("INICIO", 0)
   GraphicView "Plantilla_Visor de gráficos_1" at 80,740 size 78x6; Picture "indGris"
   GraphicView "Plantilla_Visor de gráficos_2" at 160,740 size 78x6; Picture "indGris"
   GraphicView "Plantilla_Visor de gráficos_3" at 478,740 size 78x6; Picture "indGris"
   GraphicView "Plantilla_Visor de gráficos_4" at 240,740 size 78x6; Picture "indGris"
   GraphicView "Plantilla_Visor de gráficos_5" at 557,740 size 78x6; Picture "indGris"
   GraphicView "Plantilla_Visor de gráficos_6" at 320,740 size 78x6; Picture "indGris"
   GraphicView "Plantilla_Visor de gráficos_7" at 399,740 size 78x6; Picture "indGris"
   GraphicView "Plantilla_Visor de gráficos_11" at 637,740 size 78x6; Picture "indGris"
   GraphicView "Plantilla_Visor de gráficos_8" at 80,740 size 78x6; Picture "indAmarillo"
      Visibility <- "IndCh"
   GraphicView "Plantilla_Visor de gráficos_9" at 160,740 size 78x6; Picture "indAmarillo"
      Visibility <- "IndTrCh"
   GraphicView "Plantilla_Visor de gráficos_10" at 478,740 size 78x6; Picture "indAmarillo"
      Visibility <- "IndCmpBaja"
   GraphicView "Plantilla_Visor de gráficos_12" at 240,740 size 78x6; Picture "indAmarillo"
      Visibility <- "IndCmpAlta"
   GraphicView "Plantilla_Visor de gráficos_13" at 557,740 size 78x6; Picture "indAmarillo"
      Visibility <- "IndSecBaja"
   GraphicView "Plantilla_Visor de gráficos_14" at 320,740 size 78x6; Picture "indAmarillo"
      Visibility <- "IndSecAlta"
   GraphicView "Plantilla_Visor de gráficos_15" at 399,740 size 78x6; Picture "indAmarillo"
      Visibility <- "IndTrCav"
   GraphicView "Plantilla_Visor de gráficos_16" at 637,740 size 78x6; Picture "indAmarillo"
      Visibility <- "MantenerON"
   TextField "Plantilla_Campo de texto_2" at 521,711 size 69x18; Text 'Baja Presión'
   TextField "Plantilla_Campo de texto_4" at 323,711 size 68x18; Text 'Alta Presión'
   TextField "Plantilla_Campo de texto_3" at 139,711 size 40x18; Text 'Chillers'
   Button "Plantilla_3" at 717,748 size 78x50; TextOff 'Text'; PictureOff "Rayo"
      on Click: ActivateScreen("SentronPAC-MTA", 0)
   Button "Plantilla_5" at 957,748 size 78x50; TextOff 'Text'
   Button "Plantilla_11" at 797,748 size 78x50; TextOff 'Variables Analóg.'
      on Click: ActivateScreen("Grafica", 0)
   GraphicView "Plantilla_Visor de gráficos_18" at 717,740 size 78x6; Picture "indGris"
   GraphicView "Plantilla_Visor de gráficos_19" at 797,740 size 78x6; Picture "indGris"
   GraphicView "Plantilla_Visor de gráficos_20" at 877,740 size 78x6; Picture "indGris"
   GraphicView "Plantilla_Visor de gráficos_21" at 957,740 size 78x6; Picture "indGris"
   GraphicView "Plantilla_Visor de gráficos_22" at 1037,740 size 78x6; Picture "indGris"
   GraphicView "Plantilla_Visor de gráficos_23" at 1037,740 size 78x6; Picture "indAmarillo"
      Visibility <- "AnularSirenaCav"
   Button "Plantilla_1" at 1037,749 size 78x50; TextOff 'Anular Sirena'
      on Click: SetBit("AnularSirena?")
   Button "Plantilla_2" at 1117,741 size 78x58; TextOff 'Avisos'
      on Click: ActivateScreen("MTA-Avisos", 0)
   Button "Plantilla_4" at 877,748 size 78x50; TextOff 'Text'
   GraphicView "Plantilla_Visor de gráficos_24" at 877,740 size 78x6; Picture "indGris"
   GraphicView "Plantilla_Visor de gráficos_25" at 877,740 size 78x6; Picture "indGris"
   Group "Group" at 1,716 size 1276x84
   GraphicView "Plantilla_Visor de gráficos_26" at 68,9 size 91x26; Picture "eProC logo 4 b"
   GraphicView "Plantilla_Visor de gráficos_27" at 9,8 size 49x29; Picture "eProC logo 4 a"
   GraphicView "Visor de gráficos_2" at 492,46 size 254x172; Picture "bell1"
   GraphicIOField "Plantilla_Campo ES gráfico_3" at 758,425 size 65x60; PictureList "Motor2"
      ProcessValue <- "AnimMotorMC001"
   GraphicIOField "Plantilla_Campo ES gráfico_4" at 685,353 size 65x60; PictureList "Motor2"
      ProcessValue <- "AnimMotorMC002"
   GraphicIOField "Plantilla_Campo ES gráfico_5" at 612,281 size 65x60; PictureList "Motor2"
      ProcessValue <- "AnimMotorMC004"
   GraphicIOField "Plantilla_Campo ES gráfico_2" at 539,209 size 65x60; PictureList "Motor2"
      ProcessValue <- "AnimMotorMC005"
   GraphicView "Visor de gráficos_18" at 492,46 size 254x172; Picture "Beliss2_1"
      Visibility <- "MantMC003"
   GraphicIOField "Plantilla_Campo ES gráfico_1" at 490,113 size 100x102; PictureList "MotorBelliss"
      ProcessValue <- "AnimMotorMC003"
   GraphicView "Visor de gráficos_3" at 569,134 size 246x148; Picture "ALTA1_1"
   ScreenModuleView "Faceplate_8_1" at 781,145 size 47x30
      Guid_{11997190-23981} <- "EV3"
   TextField "Plantilla_Campo de texto_1" at 1141,578 size 35x23; Text 'PT2'
   IOField "Campo ES_1" at 943,632 size 108x28; FormatPattern s999.9; Unit   bar
      ProcessValue <- "PresiónALTA"
   Button "Botón_7" at 1119,186 size 128x41; TextOff 'Tiempos'
      on Click: ActivateScreen("MTA-TiemposCmpAlta", 0)
   Button "Botón_12" at 1119,234 size 128x41; TextOff 'Presiones'
      on Click: ActivateScreen("MTA-CFGALTA", 0)
   Button "Botón_13" at 1119,138 size 128x41; TextOff 'Sopladoras'
      on Click: ActivateScreen("MTA-Sopladoras", 0)
   ScreenModuleView "Faceplate_8_5" at 927,289 size 47x30
      Guid_{11997190-23981} <- "EV4"
   ScreenModuleView "Faceplate_8_4" at 1000,361 size 47x30
      Guid_{11997190-23981} <- "EV2"
   GraphicView "Visor de gráficos_19" at 569,134 size 246x148; Picture "LOCAl"
      Visibility <- "MantMC005"
   ScreenModuleView "Faceplate_8_2" at 854,217 size 47x30
      Guid_{11997190-23981} <- "EV5"
   GraphicView "Visor de gráficos_4" at 642,206 size 246x148; Picture "ALTA1_3"
   GraphicView "Visor de gráficos_22" at 642,206 size 246x148; Picture "LOCAl"
      Visibility <- "MantMC004"
   GraphicView "Visor de gráficos_5" at 715,278 size 246x148; Picture "ALTA1_3"
   GraphicView "Visor de gráficos_21" at 715,278 size 246x148; Picture "LOCAl"
      Visibility <- "MantMC002"
   GraphicView "Visor de gráficos_6" at 788,350 size 246x148; Picture "ALTA1_3"
   GraphicView "Visor de gráficos_20" at 788,350 size 246x148; Picture "LOCAl"
      Visibility <- "MantMC001"
   ScreenModuleView "Faceplate_8_3" at 1072,433 size 47x30
      Guid_{11997190-23981} <- "EV1"
   ScreenModuleView "Faceplate_8_6" at 748,113 size 47x30
      Guid_{11997190-23981} <- "EV3b"
   ScreenModuleView "Faceplate_8_7" at 1144,505 size 47x30
      Guid_{11997190-23981} <- "EV6"
   GraphicIOField "Plantilla_Campo ES gráfico_6" at 831,497 size 65x60; PictureList "Motor2"
      ProcessValue <- "AnimMotorMC006"
   GraphicView "Visor de gráficos_1" at 861,422 size 246x148; Picture "ALTA1_3"
   GraphicView "Visor de gráficos_9" at 861,422 size 246x148; Picture "LOCAl"
      Visibility <- "MantMC006"
   Switch "Interruptor_10" at 863,114 size 40x40; TextOn '1'; TextOff '0'; CaptionText 'Switch'; PictureOff "MECH2"; Authorization "Operación"; PictureOn "MECH1"
      ProcessValue <- "MantMC003"
   Switch "Interruptor_9" at 1009,258 size 40x40; TextOn '1'; TextOff '0'; CaptionText 'Switch'; PictureOff "MECH2"; Authorization "Operación"; PictureOn "MECH1"
      ProcessValue <- "MantMC004"
   Switch "Interruptor_8" at 1082,330 size 40x40; TextOn '1'; TextOff '0'; CaptionText 'Switch'; PictureOff "MECH2"; Authorization "Operación"; PictureOn "MECH1"
      ProcessValue <- "MantMC002"
   Switch "Interruptor_6" at 936,186 size 40x40; TextOn '1'; TextOff '0'; CaptionText 'Switch'; PictureOff "MECH2"; Authorization "Operación"; PictureOn "MECH1"
      ProcessValue <- "MantMC005"
   Switch "Interruptor_7" at 1155,402 size 40x40; TextOn '1'; TextOff '0'; CaptionText 'Switch'; PictureOff "MECH2"; Authorization "Operación"; PictureOn "MECH1"
      ProcessValue <- "MantMC001"
   Switch "Interruptor_11" at 1228,474 size 40x40; TextOn '1'; TextOff '0'; CaptionText 'Switch'; PictureOff "MECH2"; Authorization "Operación"; PictureOn "MECH1"
      ProcessValue <- "MantMC006"

